(* Logix 5000 project; controller NWGG 1756-L72 rev 35.12; software revision 35.00; part 17 of 19 *)
(* tags used below, declared in another part *)
   All_Stop : BOOL;
   ALM_OVRAMP_Belt4 : ALARM_DIGITAL;
   ALM_PLUG_Belt4 : ALARM_DIGITAL;
   ALM_SLP10_Belt4 : ALARM_DIGITAL;
   ALM_SLP20_Belt4 : ALARM_DIGITAL;
   ALM_WONT_START_Belt4 : ALARM_DIGITAL;
   Auto_Start_Reversing_Belt_Fans : BOOL;
   Belt : udt_Motor[16];
   Bin_Variety_Id : STRING[30];
   Blower_707_Running : BOOL;
   Clean_Batch_Status : DINT;
   Clean_Interlock : BOOL;
   Clean_Scale_Unavailable : BOOL;
   Concrete_Leg : udt_Motor;
   ConfirmStop : BOOL;
   Current_Dist_List_IDX : DINT;
   Empty_String : STRING;
   Empty_Variety_ID : STRING;
   IDX : DINT;
   Loadout_Bin : udt_Loadout_Bin[29];
   Loadout_K_Valve : udt_Loadout_K_Valve[2];
   Longest_Treat_Start_Time : DINT;
   Longest_Treat_Stop_Time : DINT;
   Manual_Mode : BOOL;
   Manually_Start_Treater : BOOL;
   Reverse_Belt_Forward_Interlock : BOOL;
   Reverse_Belt_Stopping : BOOL;
   Reversing_Belt_Bypass_Valve : BOOL;
   Reversing_Belt_Fans : udt_Cyclone;
   Reversing_Belt_Reversed : BOOL;
   Start_Blower_707 : BOOL;
   TMR_Reverse_Delay : TIMER;
   Transfer_Batch_Status : DINT;
   Transfer_From_IDX : DINT;
   Transfer_Interlock : BOOL;
   Transfer_To_IDX : DINT;
   Treat_Batch_Status : DINT;
   Treat_Interlock : BOOL;
   Treat_Scale_Unavailable : BOOL;
   Treater_Loadout : udt_Treater_Loadout;
   Use_Concrete_Side_Clean : BOOL;
   Use_Concrete_Side_Treat : BOOL;
   Use_Steel_Side_Clean : BOOL;
   Use_Steel_Side_Treat : BOOL;
   ConcretePlantOut : DINT;
   I8_000_Bit07 : ALIAS FOR I8.7;
(* SeedLoadoutMain, continued *)

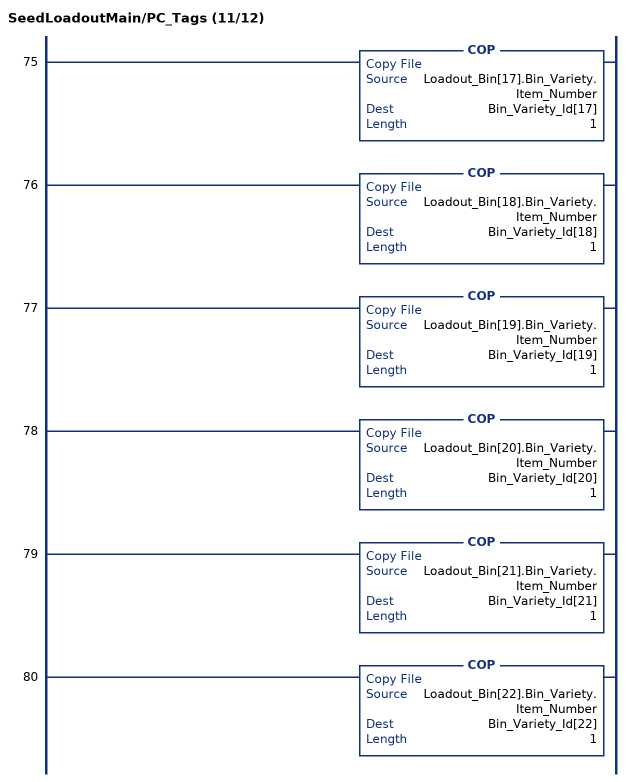
   [picture p341: SeedLoadoutMain/PC_Tags rungs 75-80]
   75: COP(Loadout_Bin[17].Bin_Variety.Item_Number,Bin_Variety_Id[17],1);
   76: COP(Loadout_Bin[18].Bin_Variety.Item_Number,Bin_Variety_Id[18],1);
   77: COP(Loadout_Bin[19].Bin_Variety.Item_Number,Bin_Variety_Id[19],1);
   78: COP(Loadout_Bin[20].Bin_Variety.Item_Number,Bin_Variety_Id[20],1);
   79: COP(Loadout_Bin[21].Bin_Variety.Item_Number,Bin_Variety_Id[21],1);
   80: COP(Loadout_Bin[22].Bin_Variety.Item_Number,Bin_Variety_Id[22],1);
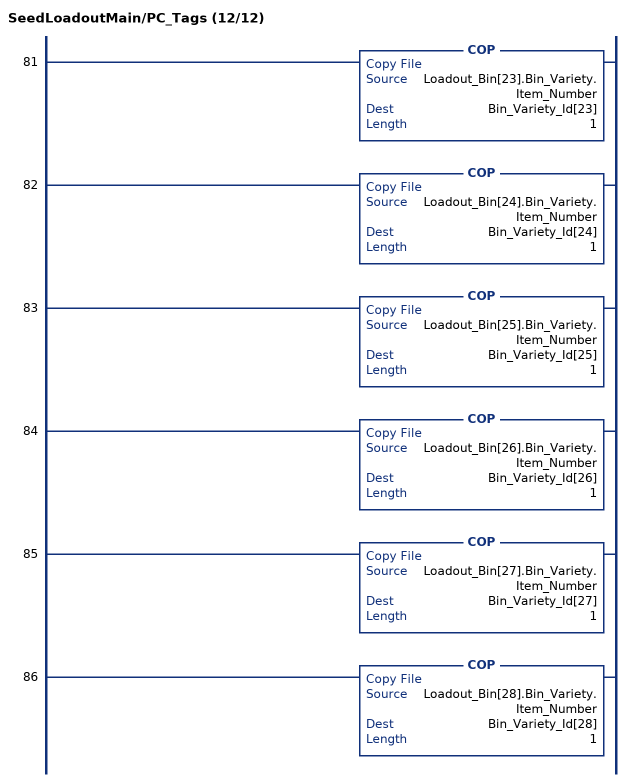
   81: COP(Loadout_Bin[23].Bin_Variety.Item_Number,Bin_Variety_Id[23],1);
   82: COP(Loadout_Bin[24].Bin_Variety.Item_Number,Bin_Variety_Id[24],1);
   83: COP(Loadout_Bin[25].Bin_Variety.Item_Number,Bin_Variety_Id[25],1);
   84: COP(Loadout_Bin[26].Bin_Variety.Item_Number,Bin_Variety_Id[26],1);
   85: COP(Loadout_Bin[27].Bin_Variety.Item_Number,Bin_Variety_Id[27],1);
   86: COP(Loadout_Bin[28].Bin_Variety.Item_Number,Bin_Variety_Id[28],1);
END_ROUTINE

ROUTINE Request_Availability   (* ladder *)
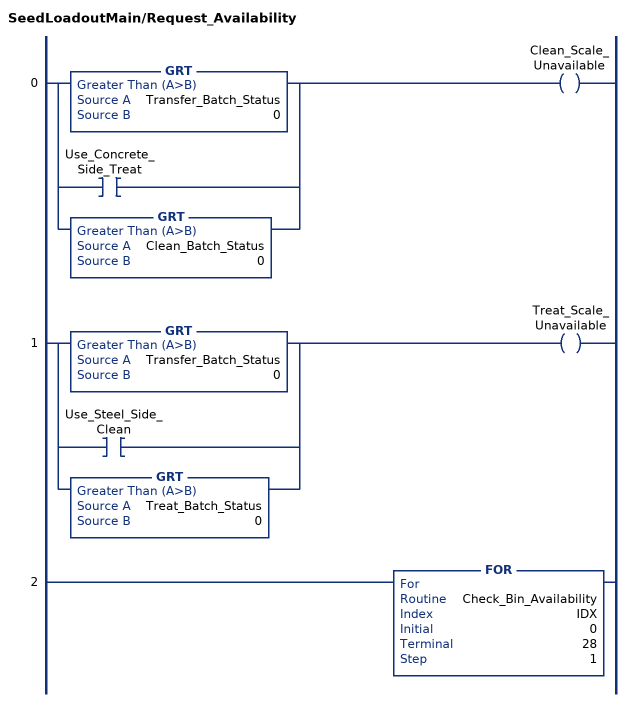
   0: [GRT(Transfer_Batch_Status,0) ,XIC(Use_Concrete_Side_Treat) ,GRT(Clean_Batch_Status,0) ]OTE(Clean_Scale_Unavailable);
   1: [GRT(Transfer_Batch_Status,0) ,XIC(Use_Steel_Side_Clean) ,GRT(Treat_Batch_Status,0) ]OTE(Treat_Scale_Unavailable);
   2: FOR(Check_Bin_Availability,IDX,0,28,1);
END_ROUTINE

ROUTINE Reset_Bin   (* ladder *)
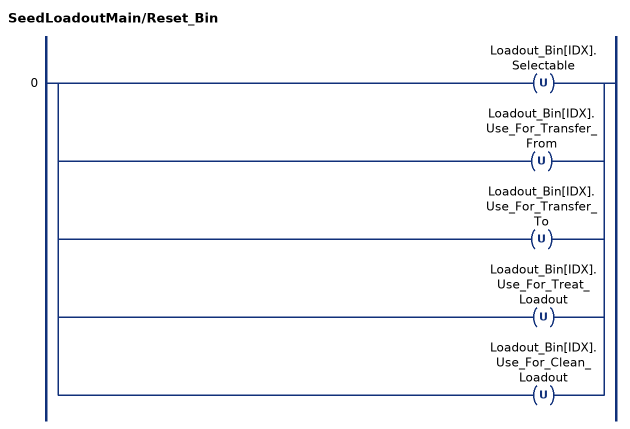
   0: [OTU(Loadout_Bin[IDX].Selectable) ,OTU(Loadout_Bin[IDX].Use_For_Transfer_From) ,OTU(Loadout_Bin[IDX].Use_For_Transfer_To) ,OTU(Loadout_Bin[IDX].Use_For_Treat_Loadout) ,OTU(Loadout_Bin[IDX].Use_For_Clean_Loadout) ];
END_ROUTINE

ROUTINE Reset_Motor_Manual   (* ladder *)
END_ROUTINE

ROUTINE Reversing_Belt   (* ladder *)
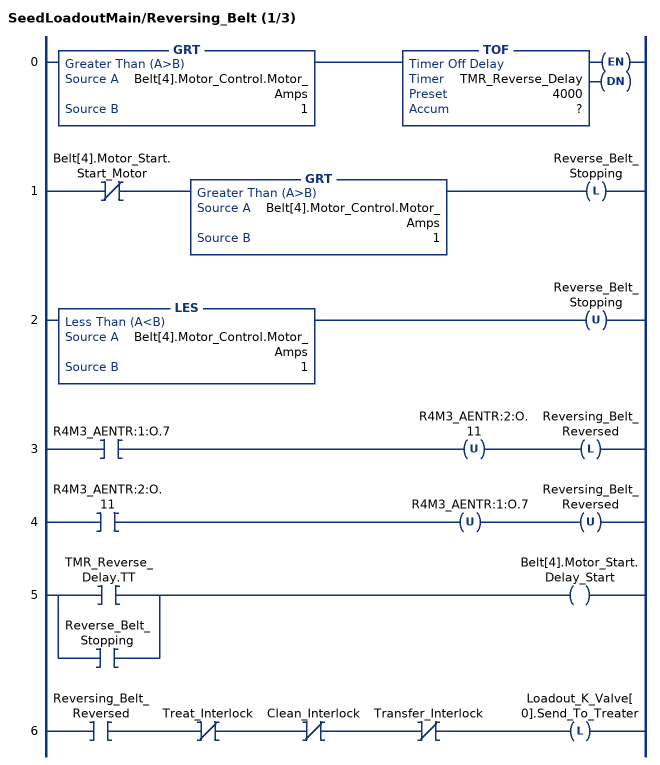
   0: GRT(Belt[4].Motor_Control.Motor_Amps,1)TOF(TMR_Reverse_Delay,?,?);
   1: XIO(Belt[4].Motor_Start.Start_Motor)GRT(Belt[4].Motor_Control.Motor_Amps,1)OTL(Reverse_Belt_Stopping);
   2: LES(Belt[4].Motor_Control.Motor_Amps,1)OTU(Reverse_Belt_Stopping);
   3: XIC(R4M3_AENTR:1:O.7)OTU(R4M3_AENTR:2:O.11)OTL(Reversing_Belt_Reversed);
   4: XIC(R4M3_AENTR:2:O.11)OTU(R4M3_AENTR:1:O.7)OTU(Reversing_Belt_Reversed);
   5: [XIC(TMR_Reverse_Delay.TT) ,XIC(Reverse_Belt_Stopping) ]OTE(Belt[4].Motor_Start.Delay_Start);
   6: XIC(Reversing_Belt_Reversed)XIO(Treat_Interlock)XIO(Clean_Interlock)XIO(Transfer_Interlock)OTL(Loadout_K_Valve[0].Send_To_Treater);
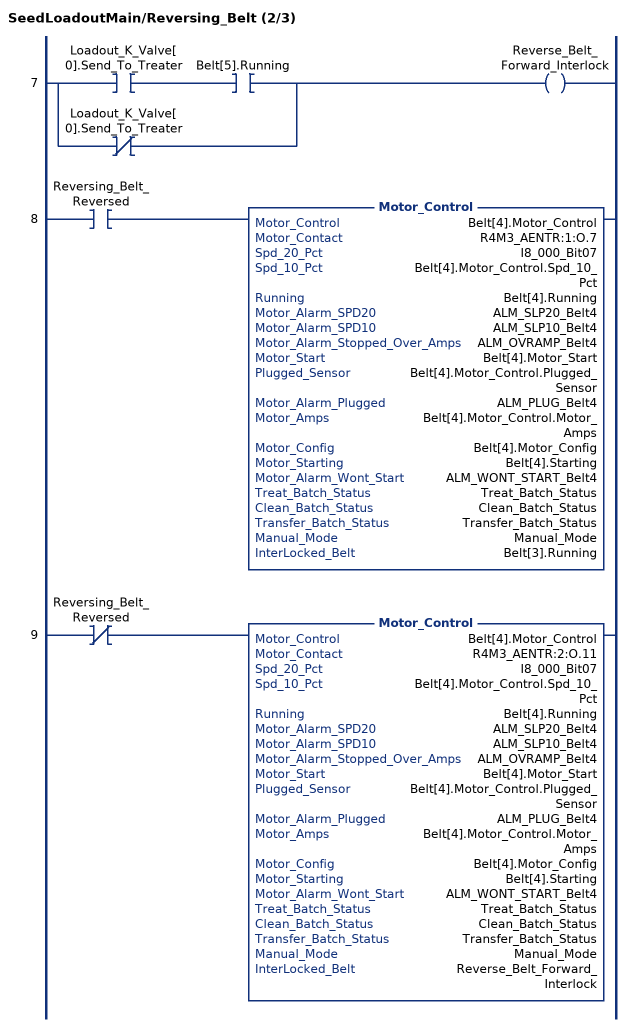
   7: [XIC(Loadout_K_Valve[0].Send_To_Treater) XIC(Belt[5].Running) ,XIO(Loadout_K_Valve[0].Send_To_Treater) ]OTE(Reverse_Belt_Forward_Interlock);
   8: XIC(Reversing_Belt_Reversed)Motor_Control(Belt[4].Motor_Control,R4M3_AENTR:1:O.7,I8_000_Bit07,Belt[4].Motor_Control.Spd_10_Pct,Belt[4].Running,ALM_SLP20_Belt4,ALM_SLP10_Belt4,ALM_OVRAMP_Belt4,Belt[4].Motor_Start,Belt[4].Motor_Control.Plugged_Sensor,ALM_PLUG_Belt4,Belt[4].Motor_Control.Motor_Amps,Belt[4].Motor_Config,Belt[4].Starting,ALM_WONT_START_Belt4,Treat_Batch_Status,Clean_Batch_Status,Transfer_Batch_Status,Manual_Mode,Belt[3].Running);
   9: XIO(Reversing_Belt_Reversed)Motor_Control(Belt[4].Motor_Control,R4M3_AENTR:2:O.11,I8_000_Bit07,Belt[4].Motor_Control.Spd_10_Pct,Belt[4].Running,ALM_SLP20_Belt4,ALM_SLP10_Belt4,ALM_OVRAMP_Belt4,Belt[4].Motor_Start,Belt[4].Motor_Control.Plugged_Sensor,ALM_PLUG_Belt4,Belt[4].Motor_Control.Motor_Amps,Belt[4].Motor_Config,Belt[4].Starting,ALM_WONT_START_Belt4,Treat_Batch_Status,Clean_Batch_Status,Transfer_Batch_Status,Manual_Mode,Reverse_Belt_Forward_Interlock);
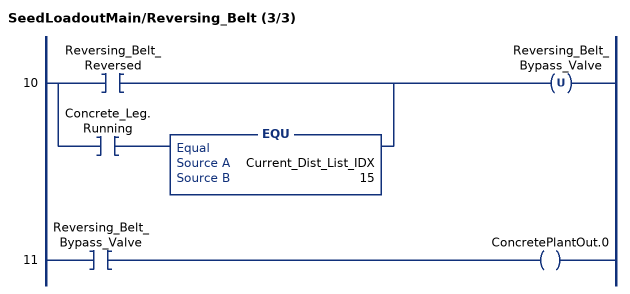
   10: [XIC(Reversing_Belt_Reversed) ,XIC(Concrete_Leg.Running) EQU(Current_Dist_List_IDX,15) ]OTU(Reversing_Belt_Bypass_Valve);
   11: XIC(Reversing_Belt_Bypass_Valve)OTE(ConcretePlantOut.0);
END_ROUTINE

ROUTINE Reversing_Belt_Fans   (* ladder *)
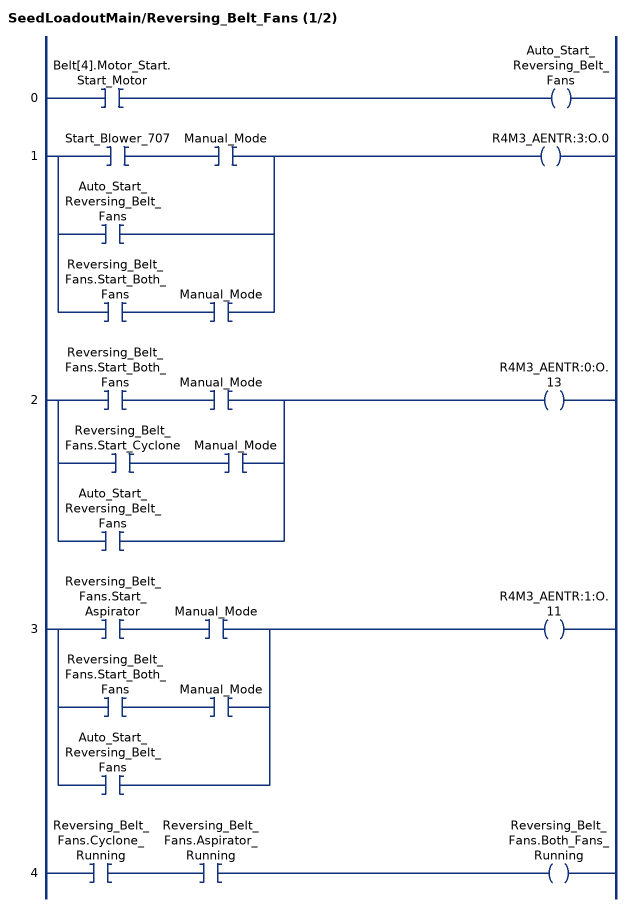
   0: XIC(Belt[4].Motor_Start.Start_Motor)OTE(Auto_Start_Reversing_Belt_Fans);
   1: [XIC(Start_Blower_707) XIC(Manual_Mode) ,XIC(Auto_Start_Reversing_Belt_Fans) ,XIC(Reversing_Belt_Fans.Start_Both_Fans) XIC(Manual_Mode) ]OTE(R4M3_AENTR:3:O.0);
   2: [XIC(Reversing_Belt_Fans.Start_Both_Fans) XIC(Manual_Mode) ,XIC(Reversing_Belt_Fans.Start_Cyclone) XIC(Manual_Mode) ,XIC(Auto_Start_Reversing_Belt_Fans) ]OTE(R4M3_AENTR:0:O.13);
   3: [XIC(Reversing_Belt_Fans.Start_Aspirator) XIC(Manual_Mode) ,XIC(Reversing_Belt_Fans.Start_Both_Fans) XIC(Manual_Mode) ,XIC(Auto_Start_Reversing_Belt_Fans) ]OTE(R4M3_AENTR:1:O.11);
   4: XIC(Reversing_Belt_Fans.Cyclone_Running)XIC(Reversing_Belt_Fans.Aspirator_Running)OTE(Reversing_Belt_Fans.Both_Fans_Running);
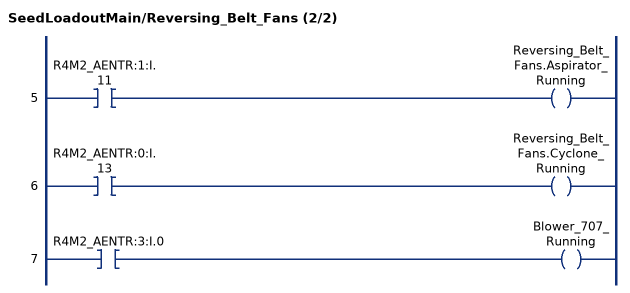
   5: XIC(R4M2_AENTR:1:I.11)OTE(Reversing_Belt_Fans.Aspirator_Running);
   6: XIC(R4M2_AENTR:0:I.13)OTE(Reversing_Belt_Fans.Cyclone_Running);
   7: XIC(R4M2_AENTR:3:I.0)OTE(Blower_707_Running);
END_ROUTINE

ROUTINE Selectable_Clean_Bins   (* ladder *)
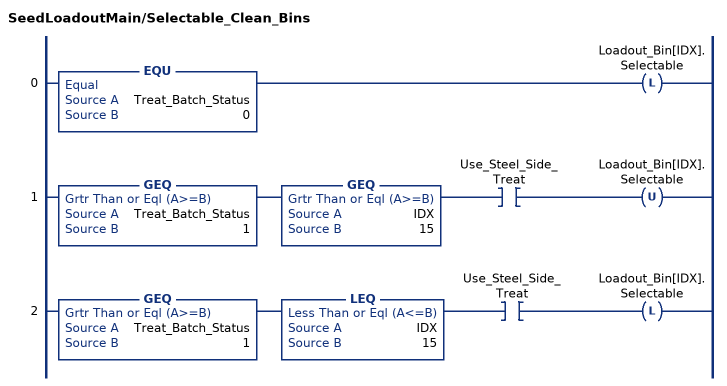
   0: EQU(Treat_Batch_Status,0)OTL(Loadout_Bin[IDX].Selectable);
   1: GEQ(Treat_Batch_Status,1)GEQ(IDX,15)XIC(Use_Steel_Side_Treat)OTU(Loadout_Bin[IDX].Selectable);
   2: GEQ(Treat_Batch_Status,1)LEQ(IDX,15)XIC(Use_Steel_Side_Treat)OTL(Loadout_Bin[IDX].Selectable);
END_ROUTINE

ROUTINE Selectable_Transfer_Bins   (* ladder *)
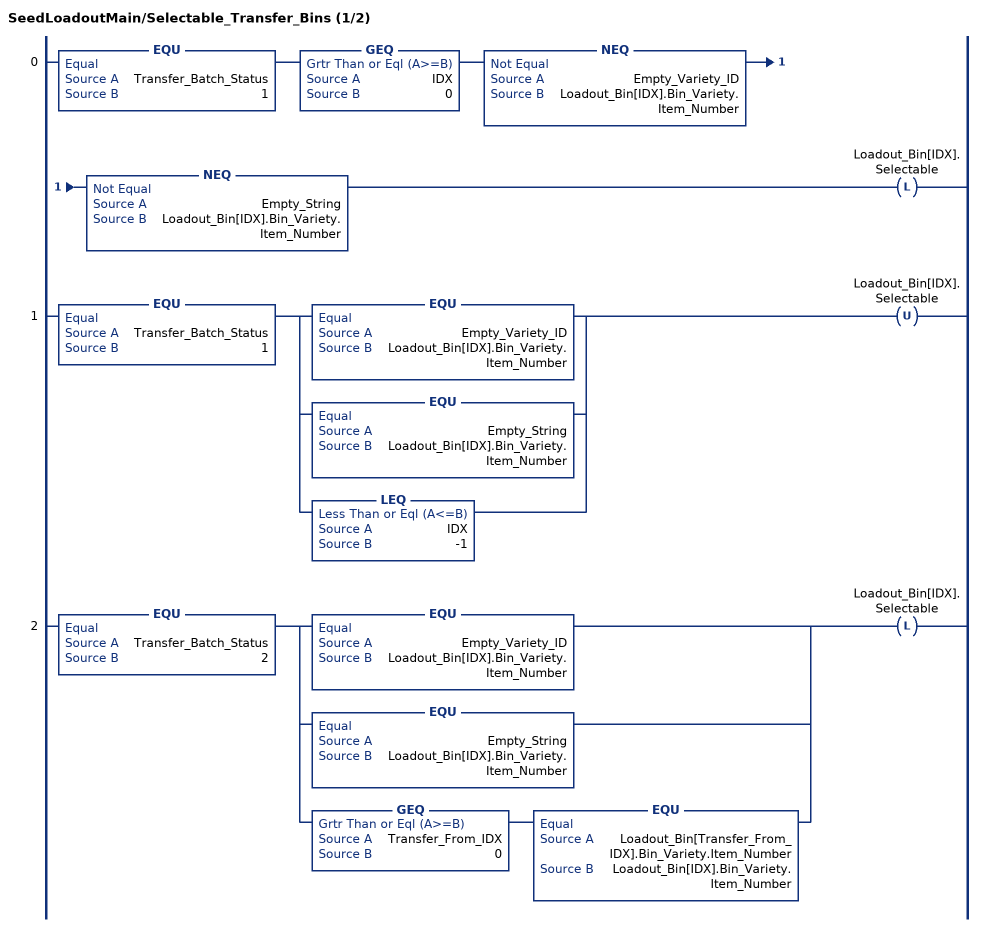
   0: EQU(Transfer_Batch_Status,1)GEQ(IDX,0)NEQ(Empty_Variety_ID,Loadout_Bin[IDX].Bin_Variety.Item_Number)NEQ(Empty_String,Loadout_Bin[IDX].Bin_Variety.Item_Number)OTL(Loadout_Bin[IDX].Selectable);
   1: EQU(Transfer_Batch_Status,1)[EQU(Empty_Variety_ID,Loadout_Bin[IDX].Bin_Variety.Item_Number) ,EQU(Empty_String,Loadout_Bin[IDX].Bin_Variety.Item_Number) ,LEQ(IDX,-1) ]OTU(Loadout_Bin[IDX].Selectable);
   2: EQU(Transfer_Batch_Status,2)[EQU(Empty_Variety_ID,Loadout_Bin[IDX].Bin_Variety.Item_Number) ,EQU(Empty_String,Loadout_Bin[IDX].Bin_Variety.Item_Number) ,GEQ(Transfer_From_IDX,0) EQU(Loadout_Bin[Transfer_From_IDX].Bin_Variety.Item_Number,Loadout_Bin[IDX].Bin_Variety.Item_Number) ]OTL(Loadout_Bin[IDX].Selectable);
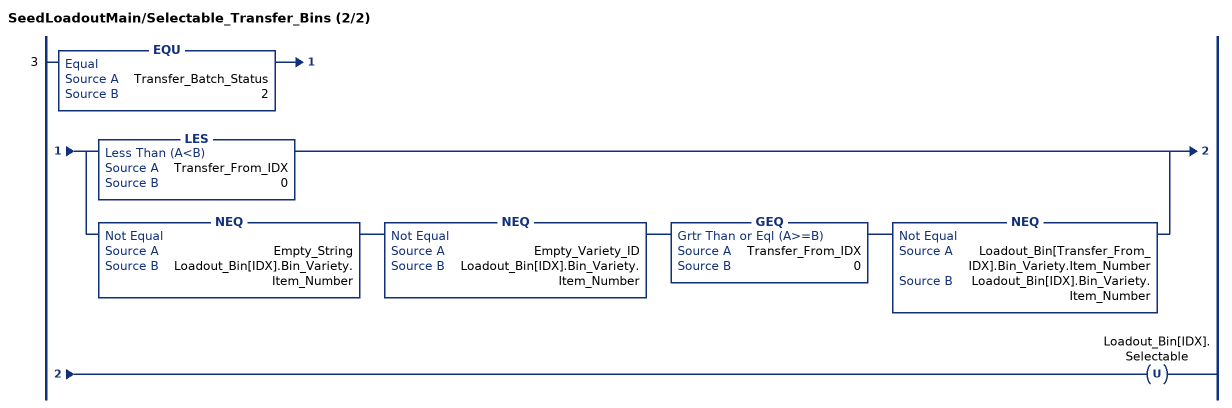
   3: EQU(Transfer_Batch_Status,2)[LES(Transfer_From_IDX,0) ,NEQ(Empty_String,Loadout_Bin[IDX].Bin_Variety.Item_Number) NEQ(Empty_Variety_ID,Loadout_Bin[IDX].Bin_Variety.Item_Number) GEQ(Transfer_From_IDX,0) NEQ(Loadout_Bin[Transfer_From_IDX].Bin_Variety.Item_Number,Loadout_Bin[IDX].Bin_Variety.Item_Number) ]OTU(Loadout_Bin[IDX].Selectable);
END_ROUTINE

ROUTINE Selectable_Treat_Bins   (* ladder *)
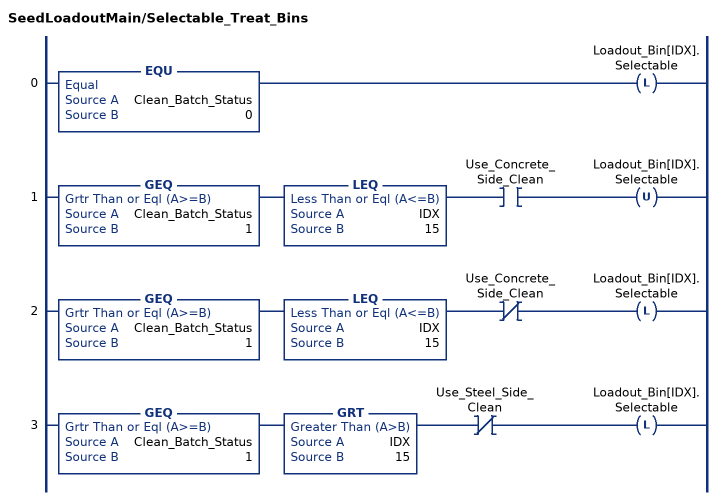
   0: EQU(Clean_Batch_Status,0)OTL(Loadout_Bin[IDX].Selectable);
   1: GEQ(Clean_Batch_Status,1)LEQ(IDX,15)XIC(Use_Concrete_Side_Clean)OTU(Loadout_Bin[IDX].Selectable);
   2: GEQ(Clean_Batch_Status,1)LEQ(IDX,15)XIO(Use_Concrete_Side_Clean)OTL(Loadout_Bin[IDX].Selectable);
   3: GEQ(Clean_Batch_Status,1)GRT(IDX,15)XIO(Use_Steel_Side_Clean)OTL(Loadout_Bin[IDX].Selectable);
END_ROUTINE

ROUTINE Set_Gate_Delay   (* ladder *)
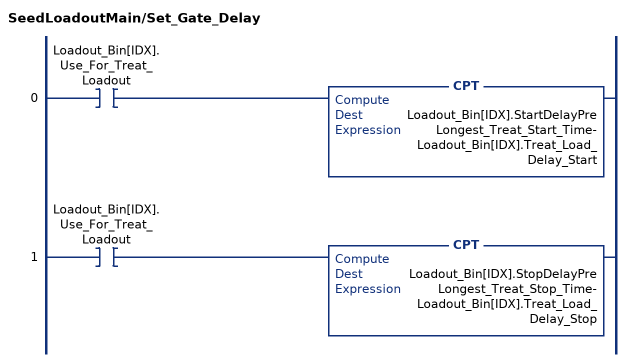
   0: XIC(Loadout_Bin[IDX].Use_For_Treat_Loadout)CPT(Loadout_Bin[IDX].StartDelayPre,Longest_Treat_Start_Time-Loadout_Bin[IDX].Treat_Load_Delay_Start);
   1: XIC(Loadout_Bin[IDX].Use_For_Treat_Loadout)CPT(Loadout_Bin[IDX].StopDelayPre,Longest_Treat_Stop_Time-Loadout_Bin[IDX].Treat_Load_Delay_Stop);
END_ROUTINE

ROUTINE Set_Transfer   (* ladder *)
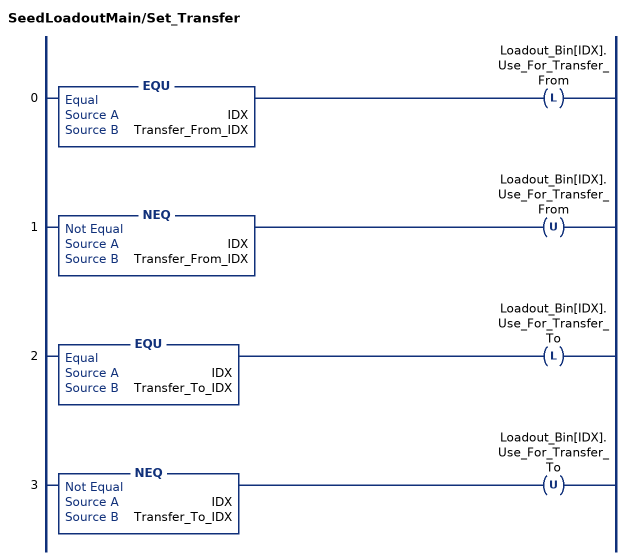
   0: EQU(IDX,Transfer_From_IDX)OTL(Loadout_Bin[IDX].Use_For_Transfer_From);
   1: NEQ(IDX,Transfer_From_IDX)OTU(Loadout_Bin[IDX].Use_For_Transfer_From);
   2: EQU(IDX,Transfer_To_IDX)OTL(Loadout_Bin[IDX].Use_For_Transfer_To);
   3: NEQ(IDX,Transfer_To_IDX)OTU(Loadout_Bin[IDX].Use_For_Transfer_To);
END_ROUTINE

ROUTINE Stop_All   (* ladder *)
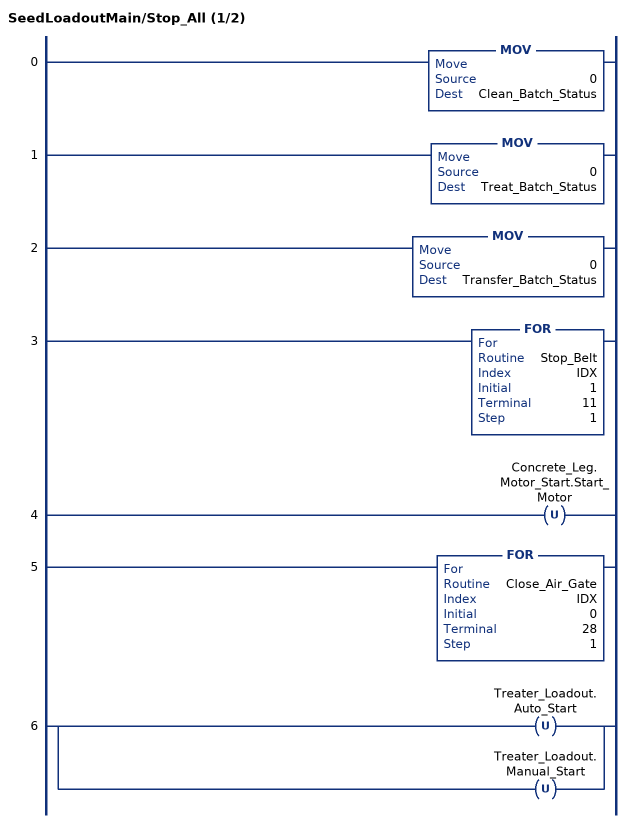
   0: MOV(0,Clean_Batch_Status);
   1: MOV(0,Treat_Batch_Status);
   2: MOV(0,Transfer_Batch_Status);
   3: FOR(Stop_Belt,IDX,1,11,1);
   4: OTU(Concrete_Leg.Motor_Start.Start_Motor);
   5: FOR(Close_Air_Gate,IDX,0,28,1);
   6: [OTU(Treater_Loadout.Auto_Start) ,OTU(Treater_Loadout.Manual_Start) ];
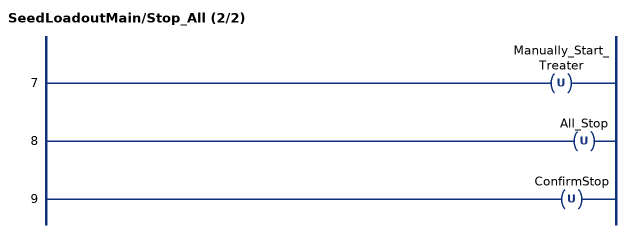
   7: OTU(Manually_Start_Treater);
   8: OTU(All_Stop);
   9: OTU(ConfirmStop);
END_ROUTINE

ROUTINE Stop_Belt   (* ladder *)
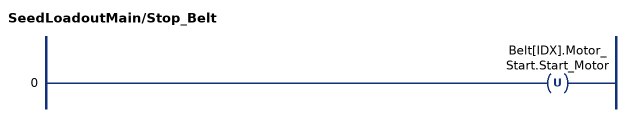
   0: OTU(Belt[IDX].Motor_Start.Start_Motor);
END_ROUTINE
